DATA_BLOCK "PanelTorreCav"   // DB21
{ S7_Optimized_Access := 'FALSE' }
VERSION : 0.1
   VAR
      InhMV030 : Bool;   // Inhibición MV030
      InhMV031 : Bool;   // Inhibición MV031
      InhMP014 : Bool;   // Inhibición MP014
      InhMP015 : Bool;   // Inhibición MP015
      Flanco1MV030 : Bool;   // Flanco 1 MV030
      Flanco1MV031 : Bool;   // Flanco 1 MV031
      Flanco1MP014 : Bool;   // Flanco 1 MP014
      Flanco1MP015 : Bool;   // Flanco 1 MP015
      Flanco2MV030 : Bool;   // Flanco 2 MV030
      Flanco2MV031 : Bool;   // Flanco 2 MV031
      Flanco2MP014 : Bool;   // Flanco 2 MP014
      Flanco2MP015 : Bool;   // Flanco 2 MP015
      Flanco3MV030 : Bool;   // Flanco 3 MV030
      Flanco3MV031 : Bool;   // Flanco 3 MV031
      Flanco3MP014 : Bool;   // Flanco 3 MP014
      Flanco3MP015 : Bool;   // Flanco 3 MP015
      HabPanelMV030 : Bool;   // Habilitación desde Panel MV030
      HabPanelMV031 : Bool;   // Habilitación desde Panel MV031
      HabPanelMP014 : Bool;   // Habilitación desde Panel MP014
      HabPanelMP015 : Bool;   // Habilitación desde Panel MP015
      DeshabPanelMV030 : Bool;   // Deshabilitación desde Panel MV030
      DeshabPanelMV031 : Bool;   // Deshabilitación desde Panel MV031
      DeshabPanelMP014 : Bool;   // Deshabilitación desde Panel MP014
      DeshabPanelMP015 : Bool;   // Deshabilitación desde Panel MP015
      MarchaPanelMV030 : Bool;   // Marcha desde Panel MV030
      MarchaPanelMV031 : Bool;   // Marcha desde Panel MV031
      MarchaPanelMP014 : Bool;   // Marcha desde Panel MP014
      MarchaPanelMP015 : Bool;   // Marcha desde Panel MP015
      ParadaPanelMV030 : Bool;   // Parada desde Panel MV030
      ParadaPanelMV031 : Bool;   // Parada desde Panel MV031
      ParadaPanelMP014 : Bool;   // Parada desde Panel MP014
      ParadaPanelMP015 : Bool;   // Parada desde Panel MP015
      HabMV030 : Bool;   // Habilitado MV030
      HabMV031 : Bool;   // Habilitado MV031
      HabMP014 : Bool;   // Habilitado MP014
      HabMP015 : Bool;   // Habilitado MP015
      DeshabMV030 : Bool;   // Deshabilitado MV030
      DeshabMV031 : Bool;   // Deshabilitado MV031
      DeshabMP014 : Bool;   // Deshabilitado MP014
      DeshabMP015 : Bool;   // Deshabilitado MP015
      MarchaMV030 : Bool;   // Marchando MV030
      MarchaMV031 : Bool;   // Marchando MV031
      MarchaMP014 : Bool;   // Marchando MP014
      MarchaMP015 : Bool;   // Marchando MP015
      ParadaMV030 : Bool;   // Parando MV030
      ParadaMV031 : Bool;   // Parando MV031
      ParadaMP014 : Bool;   // Parando MP014
      ParadaMP015 : Bool;   // Parando MP015
      MantMV030 : Bool;   // Mantenimiento MV030
      MantMV031 : Bool;   // Mantenimiento MV031
      MantMP014 : Bool;   // Mantenimiento MP014
      MantMP015 : Bool;   // Mantenimiento MP015
      AutoV030 : Bool;   // Ventilador Controlado por temperatura V030
      AutoV031 : Bool;   // Ventilador Controlado por temperatura V031
      SPonV030 : Int;   // Setpoint arranque para V001
      SPonV031 : Int;   // Setpoint arranque para V002
      SPoffV030 : Int;   // Setpoint parada para V001
      SPoffV031 : Int;   // Setpoint parada para V002
      Temperatura : Int;   // Temperatura agua de torres
      ArranqueAutoV030 : Bool;   // Arranque Automático de ventilador 1
      ArranqueAutoV031 : Bool;   // Arranque Automático de ventilador 2
      Reserva_13 : Bool;
      Reserva_14 : Bool;
      Reserva_15 : Bool;
      Reserva_16 : Bool;
      Reserva_17 : Bool;
      Reserva_18 : Bool;
      Reserva_19 : Bool;
      Reserva_110 : Bool;
      Reserva_111 : Bool;
      Reserva_112 : Bool;
      Reserva_113 : Bool;
      Reserva_114 : Bool;
      Reserva_115 : Bool;
      Reserva_116 : Bool;
      Reserva_117 : Bool;
      Reserva_118 : Bool;
      Reserva_119 : Bool;
      Reserva_120 : Bool;
      Reserva_121 : Bool;
      Reserva_122 : Bool;
      Reserva_123 : Bool;
      Reserva_124 : Bool;
      Reserva_125 : Bool;
      Reserva_126 : Bool;
      Reserva_127 : Bool;
      Reserva_128 : Bool;
      Reserva_129 : Bool;
      Reserva_130 : Bool;
      Reserva_131 : Bool;
      Reserva_132 : Bool;
      Reserva_133 : Bool;
      Reserva_134 : Bool;
      Reserva_135 : Bool;
      Reserva_136 : Bool;
      Reserva_137 : Bool;
      Reserva_138 : Bool;
      Reserva_139 : Bool;
      Reserva_140 : Bool;
      Reserva_141 : Bool;
      Reserva_142 : Bool;
      Reserva_143 : Bool;
   END_VAR
BEGIN
END_DATA_BLOCK

DATA_BLOCK "TAguaCAV"   // DB51
{ S7_Optimized_Access := 'FALSE' }
AUTHOR : AEB
VERSION : 0.1
   VAR
      PrAlta : Real := 3.585069e+1;   // Presión Aire de Alta
      TmpCav : Real := 2.061632e+1;   // Temp Torre Cavaleto
      PrAlta2 : Real := 3.541667e+1;   // Presión Aire de Alta_Redundante
      PrBaja : Real := 6.140046e+0;   // Presión Aire de Baja
      STAT4 : Real;
      STAT5 : Real;
      STAT6 : Real;
      STAT7 : Real;
      STAT8 : Real;
      STAT9 : Real;
      STAT10 : Real := 1.446759e-3;
      STAT11 : Real;
      STAT12 : Real;
      STAT13 : Real;
      STAT14 : Real;
      STAT15 : Real;
      STAT16 : Real;
      STAT17 : Real;
      STAT18 : Real;
      STAT19 : Real;
      STAT20 : Real;
      STAT21 : Real;
      STAT22 : Real;
      STAT23 : Real;
      STAT24 : Real;
      STAT25 : Real;
      STAT26 : Real;
      STAT27 : Real;
      STAT28 : Real;
      STAT29 : Real;
      STAT30 : Real;
      STAT31 : Real;
      STAT32 : Real;
      STAT33 : Real;
      STAT34 : Real;
      STAT35 : Real;
      STAT36 : Real;
      STAT37 : Real;
      STAT38 : Real;
      STAT39 : Real;
      STAT40 : Real;
      STAT41 : Real;
      STAT42 : Real;
      STAT43 : Real;
      STAT44 : Real;
      STAT45 : Real;
      STAT46 : Real;
      STAT47 : Real;
      STAT48 : Real;
      STAT49 : Real;
      STAT50 : Real;
      STAT51 : Real;
      STAT52 : Real;
      STAT53 : Real;
      STAT54 : Real;
      STAT55 : Real;
      STAT56 : Real;
      STAT57 : Real;
      STAT58 : Real;
      STAT59 : Real;
      STAT60 : Real;
      STAT61 : Real;
      STAT62 : Real;
      STAT63 : Real;
      STAT64 : Real;
      STAT65 : Real;
   END_VAR
BEGIN
END_DATA_BLOCK

// folder: Torres de Agua/Torres Chillers

DATA_BLOCK "CFG-TorresCH"   // DB92
{ S7_Optimized_Access := 'FALSE' }
VERSION : 0.1
   VAR
      AutoV001 : Bool;   // Ventilador Controlado por temperatura V001
      AutoV002 : Bool;   // Ventilador Controlado por temperatura V002
      AutoV003 : Bool;   // Ventilador Controlado por temperatura V003
      SPonV001 : Int;   // Setpoint arranque para V001
      SPonV002 : Int;   // Setpoint arranque para V002
      SPonV003 : Int;   // Setpoint arranque para V003
      SPoffV001 : Int;   // Setpoint parada para V001
      SPoffV002 : Int;   // Setpoint parada para V002
      SPoffV003 : Int;   // Setpoint parada para V003
      Temperatura : Int;   // Temperatura agua de torres
      ArranqueAutoV001 : Bool;   // Arranque Automático de ventilador 1
      ArranqueAutoV002 : Bool;   // Arranque Automático de ventilador 2
      ArranqueAutoV003 : Bool;   // Arranque Automático de ventilador 3
   END_VAR
BEGIN
END_DATA_BLOCK

// folder: (top level)

FUNCTION "Arranques General" : Void   // FC4, LAD
{ S7_Optimized_Access := 'FALSE' }
VERSION : 0.1
   VAR_TEMP
      TEMP0 : Bool;
      TEMP1 : Bool;
      TEMP2 : Bool;
      TEMP3 : Bool;
      TEMP4 : Bool;
   END_VAR
   VAR_TEMP   // added for the SCL form of the ladder/FBD networks
      _w1 : Bool;
      _w2 : Bool;
      _s5time1 : S5Time;
   END_VAR
BEGIN

REGION Network 1: Motor MT007 - Bomba Soplado L1 / Bloque motor MT007 - Bomba Soplado L1
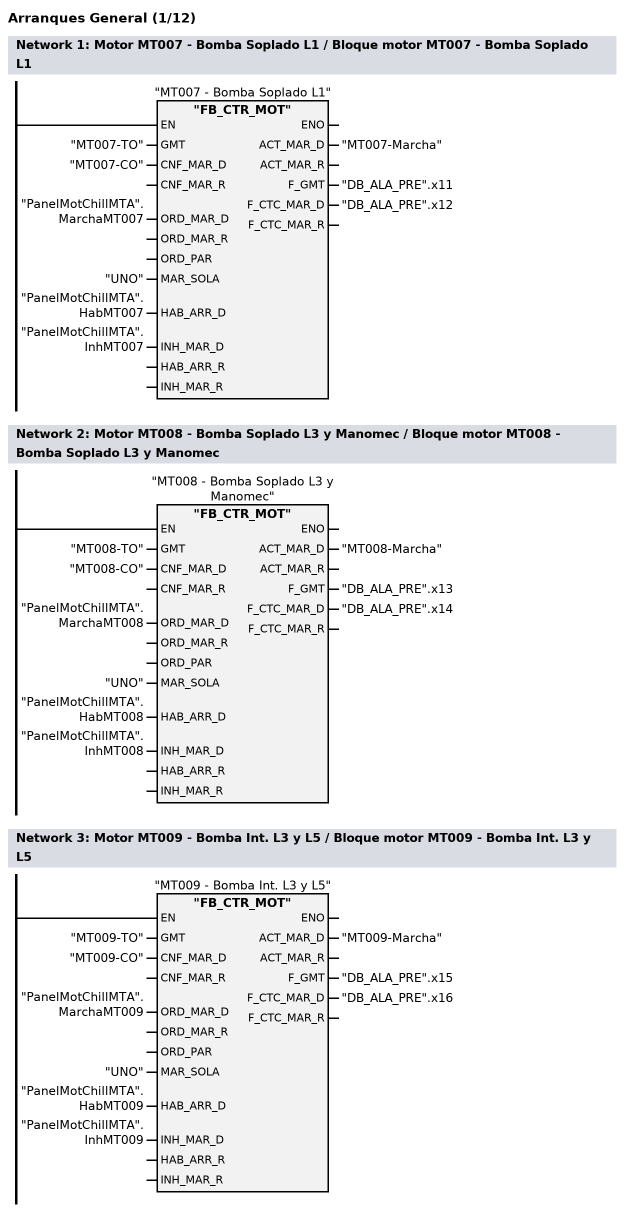
   RUNG wire#powerrail
      "MT007 - Bomba Soplado L1"(GMT := "MT007-TO", CNF_MAR_D := "MT007-CO", CNF_MAR_R :=, ORD_MAR_D := "PanelMotChillMTA".MarchaMT007, ORD_MAR_R :=, ORD_PAR :=, MAR_SOLA := "UNO", HAB_ARR_D := "PanelMotChillMTA".HabMT007, INH_MAR_D := "PanelMotChillMTA".InhMT007, HAB_ARR_R :=, INH_MAR_R :=, ACT_MAR_D => "MT007-Marcha", ACT_MAR_R =>, F_GMT => "DB_ALA_PRE".x11, F_CTC_MAR_D => "DB_ALA_PRE".x12, F_CTC_MAR_R =>)
   END_RUNG
   // the same network as SCL:
   "MT007 - Bomba Soplado L1"(GMT := "MT007-TO",   // "FB_CTR_MOT"
                           CNF_MAR_D := "MT007-CO",
                           ORD_MAR_D := "PanelMotChillMTA".MarchaMT007,
                           MAR_SOLA := "UNO",
                           HAB_ARR_D := "PanelMotChillMTA".HabMT007,
                           INH_MAR_D := "PanelMotChillMTA".InhMT007,
                           ACT_MAR_D => "MT007-Marcha",
                           F_GMT => "DB_ALA_PRE".x11,
                           F_CTC_MAR_D => "DB_ALA_PRE".x12);
END_REGION

REGION Network 2: Motor MT008 - Bomba Soplado L3 y Manomec / Bloque motor MT008 - Bomba Soplado L3 y Manomec
   RUNG wire#powerrail
      "MT008 - Bomba Soplado L3 y Manomec"(GMT := "MT008-TO", CNF_MAR_D := "MT008-CO", CNF_MAR_R :=, ORD_MAR_D := "PanelMotChillMTA".MarchaMT008, ORD_MAR_R :=, ORD_PAR :=, MAR_SOLA := "UNO", HAB_ARR_D := "PanelMotChillMTA".HabMT008, INH_MAR_D := "PanelMotChillMTA".InhMT008, HAB_ARR_R :=, INH_MAR_R :=, ACT_MAR_D => "MT008-Marcha", ACT_MAR_R =>, F_GMT => "DB_ALA_PRE".x13, F_CTC_MAR_D => "DB_ALA_PRE".x14, F_CTC_MAR_R =>)
   END_RUNG
   // the same network as SCL:
   "MT008 - Bomba Soplado L3 y Manomec"(GMT := "MT008-TO",   // "FB_CTR_MOT"
                           CNF_MAR_D := "MT008-CO",
                           ORD_MAR_D := "PanelMotChillMTA".MarchaMT008,
                           MAR_SOLA := "UNO",
                           HAB_ARR_D := "PanelMotChillMTA".HabMT008,
                           INH_MAR_D := "PanelMotChillMTA".InhMT008,
                           ACT_MAR_D => "MT008-Marcha",
                           F_GMT => "DB_ALA_PRE".x13,
                           F_CTC_MAR_D => "DB_ALA_PRE".x14);
END_REGION

REGION Network 3: Motor MT009 - Bomba Int. L3 y L5 / Bloque motor MT009 - Bomba Int. L3 y L5
   RUNG wire#powerrail
      "MT009 - Bomba Int. L3 y L5"(GMT := "MT009-TO", CNF_MAR_D := "MT009-CO", CNF_MAR_R :=, ORD_MAR_D := "PanelMotChillMTA".MarchaMT009, ORD_MAR_R :=, ORD_PAR :=, MAR_SOLA := "UNO", HAB_ARR_D := "PanelMotChillMTA".HabMT009, INH_MAR_D := "PanelMotChillMTA".InhMT009, HAB_ARR_R :=, INH_MAR_R :=, ACT_MAR_D => "MT009-Marcha", ACT_MAR_R =>, F_GMT => "DB_ALA_PRE".x15, F_CTC_MAR_D => "DB_ALA_PRE".x16, F_CTC_MAR_R =>)
   END_RUNG
   // the same network as SCL:
   "MT009 - Bomba Int. L3 y L5"(GMT := "MT009-TO",   // "FB_CTR_MOT"
                           CNF_MAR_D := "MT009-CO",
                           ORD_MAR_D := "PanelMotChillMTA".MarchaMT009,
                           MAR_SOLA := "UNO",
                           HAB_ARR_D := "PanelMotChillMTA".HabMT009,
                           INH_MAR_D := "PanelMotChillMTA".InhMT009,
                           ACT_MAR_D => "MT009-Marcha",
                           F_GMT => "DB_ALA_PRE".x15,
                           F_CTC_MAR_D => "DB_ALA_PRE".x16);
END_REGION

REGION Network 4: Motor MT010 - Bomba Int L1 y Manomec / Bloque motor MT010 - Bomba Int L1 y Manomec
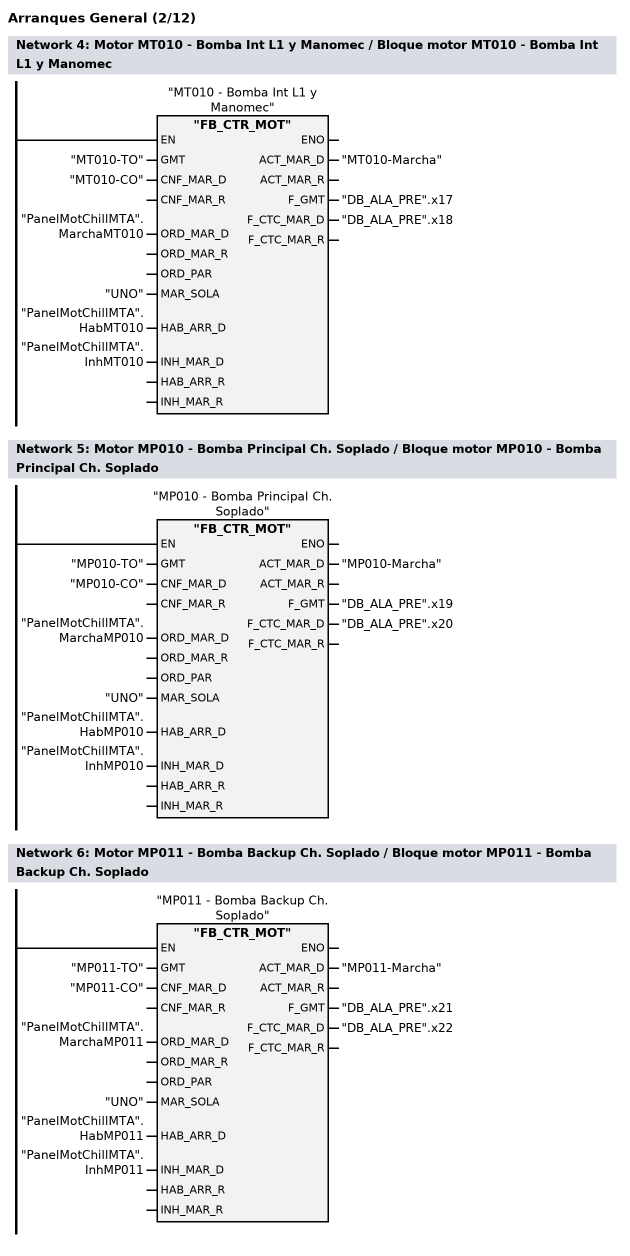
   RUNG wire#powerrail
      "MT010 - Bomba Int L1 y Manomec"(GMT := "MT010-TO", CNF_MAR_D := "MT010-CO", CNF_MAR_R :=, ORD_MAR_D := "PanelMotChillMTA".MarchaMT010, ORD_MAR_R :=, ORD_PAR :=, MAR_SOLA := "UNO", HAB_ARR_D := "PanelMotChillMTA".HabMT010, INH_MAR_D := "PanelMotChillMTA".InhMT010, HAB_ARR_R :=, INH_MAR_R :=, ACT_MAR_D => "MT010-Marcha", ACT_MAR_R =>, F_GMT => "DB_ALA_PRE".x17, F_CTC_MAR_D => "DB_ALA_PRE".x18, F_CTC_MAR_R =>)
   END_RUNG
   // the same network as SCL:
   "MT010 - Bomba Int L1 y Manomec"(GMT := "MT010-TO",   // "FB_CTR_MOT"
                           CNF_MAR_D := "MT010-CO",
                           ORD_MAR_D := "PanelMotChillMTA".MarchaMT010,
                           MAR_SOLA := "UNO",
                           HAB_ARR_D := "PanelMotChillMTA".HabMT010,
                           INH_MAR_D := "PanelMotChillMTA".InhMT010,
                           ACT_MAR_D => "MT010-Marcha",
                           F_GMT => "DB_ALA_PRE".x17,
                           F_CTC_MAR_D => "DB_ALA_PRE".x18);
END_REGION

REGION Network 5: Motor MP010 - Bomba Principal Ch. Soplado / Bloque motor MP010 - Bomba Principal Ch. Soplado
   RUNG wire#powerrail
      "MP010 - Bomba Principal Ch. Soplado"(GMT := "MP010-TO", CNF_MAR_D := "MP010-CO", CNF_MAR_R :=, ORD_MAR_D := "PanelMotChillMTA".MarchaMP010, ORD_MAR_R :=, ORD_PAR :=, MAR_SOLA := "UNO", HAB_ARR_D := "PanelMotChillMTA".HabMP010, INH_MAR_D := "PanelMotChillMTA".InhMP010, HAB_ARR_R :=, INH_MAR_R :=, ACT_MAR_D => "MP010-Marcha", ACT_MAR_R =>, F_GMT => "DB_ALA_PRE".x19, F_CTC_MAR_D => "DB_ALA_PRE".x20, F_CTC_MAR_R =>)
   END_RUNG
   // the same network as SCL:
   "MP010 - Bomba Principal Ch. Soplado"(GMT := "MP010-TO",   // "FB_CTR_MOT"
                           CNF_MAR_D := "MP010-CO",
                           ORD_MAR_D := "PanelMotChillMTA".MarchaMP010,
                           MAR_SOLA := "UNO",
                           HAB_ARR_D := "PanelMotChillMTA".HabMP010,
                           INH_MAR_D := "PanelMotChillMTA".InhMP010,
                           ACT_MAR_D => "MP010-Marcha",
                           F_GMT => "DB_ALA_PRE".x19,
                           F_CTC_MAR_D => "DB_ALA_PRE".x20);
END_REGION

REGION Network 6: Motor MP011 - Bomba Backup Ch. Soplado / Bloque motor MP011 - Bomba Backup Ch. Soplado
   RUNG wire#powerrail
      "MP011 - Bomba Backup Ch. Soplado"(GMT := "MP011-TO", CNF_MAR_D := "MP011-CO", CNF_MAR_R :=, ORD_MAR_D := "PanelMotChillMTA".MarchaMP011, ORD_MAR_R :=, ORD_PAR :=, MAR_SOLA := "UNO", HAB_ARR_D := "PanelMotChillMTA".HabMP011, INH_MAR_D := "PanelMotChillMTA".InhMP011, HAB_ARR_R :=, INH_MAR_R :=, ACT_MAR_D => "MP011-Marcha", ACT_MAR_R =>, F_GMT => "DB_ALA_PRE".x21, F_CTC_MAR_D => "DB_ALA_PRE".x22, F_CTC_MAR_R =>)
   END_RUNG
   // the same network as SCL:
   "MP011 - Bomba Backup Ch. Soplado"(GMT := "MP011-TO",   // "FB_CTR_MOT"
                           CNF_MAR_D := "MP011-CO",
                           ORD_MAR_D := "PanelMotChillMTA".MarchaMP011,
                           MAR_SOLA := "UNO",
                           HAB_ARR_D := "PanelMotChillMTA".HabMP011,
                           INH_MAR_D := "PanelMotChillMTA".InhMP011,
                           ACT_MAR_D => "MP011-Marcha",
                           F_GMT => "DB_ALA_PRE".x21,
                           F_CTC_MAR_D => "DB_ALA_PRE".x22);
END_REGION

REGION Network 7: Motor MP012 - Bomba Principal Ch. Envasado / Bloque motor MP012 - Bomba Principal Ch. Envasado
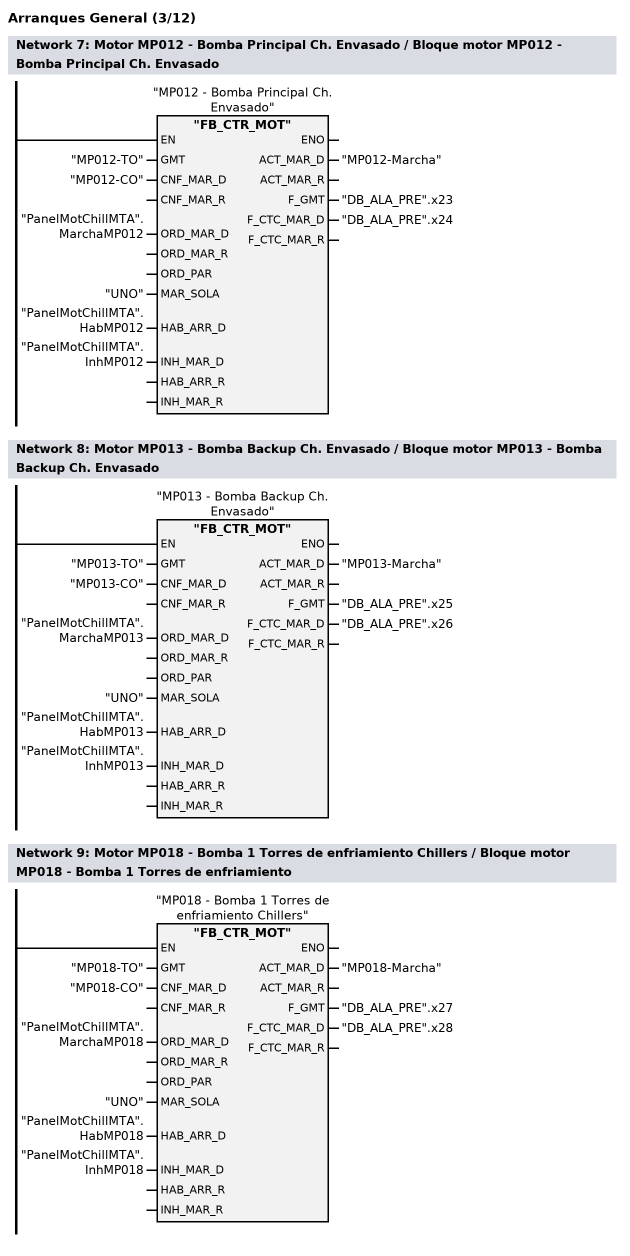
   RUNG wire#powerrail
      "MP012 - Bomba Principal Ch. Envasado"(GMT := "MP012-TO", CNF_MAR_D := "MP012-CO", CNF_MAR_R :=, ORD_MAR_D := "PanelMotChillMTA".MarchaMP012, ORD_MAR_R :=, ORD_PAR :=, MAR_SOLA := "UNO", HAB_ARR_D := "PanelMotChillMTA".HabMP012, INH_MAR_D := "PanelMotChillMTA".InhMP012, HAB_ARR_R :=, INH_MAR_R :=, ACT_MAR_D => "MP012-Marcha", ACT_MAR_R =>, F_GMT => "DB_ALA_PRE".x23, F_CTC_MAR_D => "DB_ALA_PRE".x24, F_CTC_MAR_R =>)
   END_RUNG
   // the same network as SCL:
   "MP012 - Bomba Principal Ch. Envasado"(GMT := "MP012-TO",   // "FB_CTR_MOT"
                           CNF_MAR_D := "MP012-CO",
                           ORD_MAR_D := "PanelMotChillMTA".MarchaMP012,
                           MAR_SOLA := "UNO",
                           HAB_ARR_D := "PanelMotChillMTA".HabMP012,
                           INH_MAR_D := "PanelMotChillMTA".InhMP012,
                           ACT_MAR_D => "MP012-Marcha",
                           F_GMT => "DB_ALA_PRE".x23,
                           F_CTC_MAR_D => "DB_ALA_PRE".x24);
END_REGION

REGION Network 8: Motor MP013 - Bomba Backup Ch. Envasado / Bloque motor MP013 - Bomba Backup Ch. Envasado
   RUNG wire#powerrail
      "MP013 - Bomba Backup Ch. Envasado"(GMT := "MP013-TO", CNF_MAR_D := "MP013-CO", CNF_MAR_R :=, ORD_MAR_D := "PanelMotChillMTA".MarchaMP013, ORD_MAR_R :=, ORD_PAR :=, MAR_SOLA := "UNO", HAB_ARR_D := "PanelMotChillMTA".HabMP013, INH_MAR_D := "PanelMotChillMTA".InhMP013, HAB_ARR_R :=, INH_MAR_R :=, ACT_MAR_D => "MP013-Marcha", ACT_MAR_R =>, F_GMT => "DB_ALA_PRE".x25, F_CTC_MAR_D => "DB_ALA_PRE".x26, F_CTC_MAR_R =>)
   END_RUNG
   // the same network as SCL:
   "MP013 - Bomba Backup Ch. Envasado"(GMT := "MP013-TO",   // "FB_CTR_MOT"
                           CNF_MAR_D := "MP013-CO",
                           ORD_MAR_D := "PanelMotChillMTA".MarchaMP013,
                           MAR_SOLA := "UNO",
                           HAB_ARR_D := "PanelMotChillMTA".HabMP013,
                           INH_MAR_D := "PanelMotChillMTA".InhMP013,
                           ACT_MAR_D => "MP013-Marcha",
                           F_GMT => "DB_ALA_PRE".x25,
                           F_CTC_MAR_D => "DB_ALA_PRE".x26);
END_REGION

REGION Network 9: Motor MP018 - Bomba 1 Torres de enfriamiento Chillers / Bloque motor MP018 - Bomba 1 Torres de enfriamiento
   RUNG wire#powerrail
      "MP018 - Bomba 1 Torres de enfriamiento Chillers"(GMT := "MP018-TO", CNF_MAR_D := "MP018-CO", CNF_MAR_R :=, ORD_MAR_D := "PanelMotChillMTA".MarchaMP018, ORD_MAR_R :=, ORD_PAR :=, MAR_SOLA := "UNO", HAB_ARR_D := "PanelMotChillMTA".HabMP018, INH_MAR_D := "PanelMotChillMTA".InhMP018, HAB_ARR_R :=, INH_MAR_R :=, ACT_MAR_D => "MP018-Marcha", ACT_MAR_R =>, F_GMT => "DB_ALA_PRE".x27, F_CTC_MAR_D => "DB_ALA_PRE".x28, F_CTC_MAR_R =>)
   END_RUNG
   // the same network as SCL:
   "MP018 - Bomba 1 Torres de enfriamiento Chillers"(GMT := "MP018-TO",   // "FB_CTR_MOT"
                           CNF_MAR_D := "MP018-CO",
                           ORD_MAR_D := "PanelMotChillMTA".MarchaMP018,
                           MAR_SOLA := "UNO",
                           HAB_ARR_D := "PanelMotChillMTA".HabMP018,
                           INH_MAR_D := "PanelMotChillMTA".InhMP018,
                           ACT_MAR_D => "MP018-Marcha",
                           F_GMT => "DB_ALA_PRE".x27,
                           F_CTC_MAR_D => "DB_ALA_PRE".x28);
END_REGION

REGION Network 10: Motor MP019 - Bomba 2 Torres de enfriamiento Chillers / Bloque motor MP019 - Bomba 2 Torres de enfriamiento
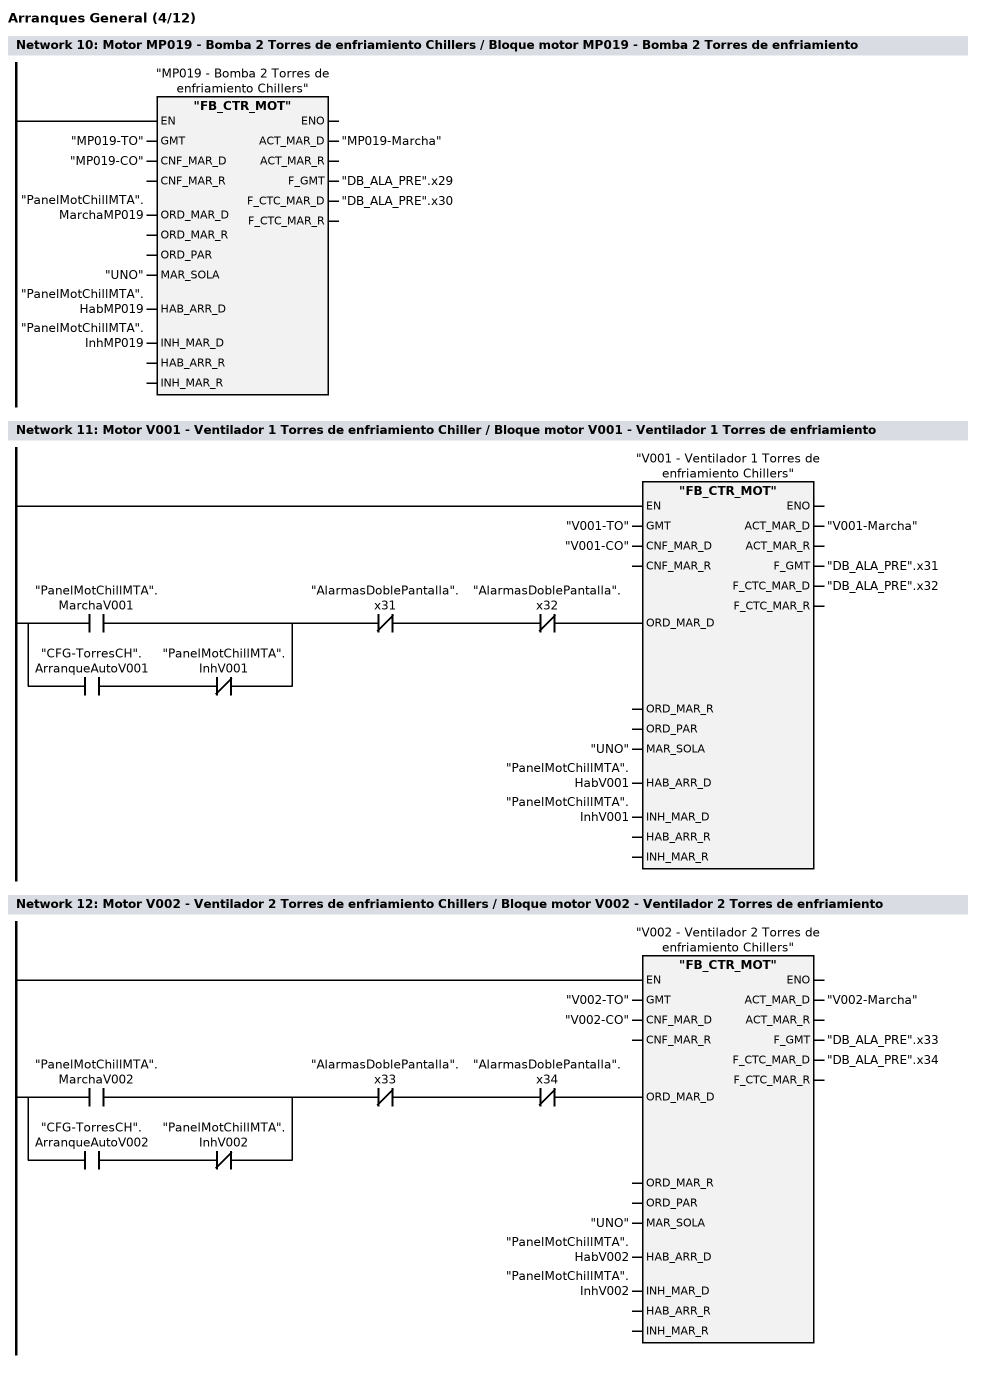
   RUNG wire#powerrail
      "MP019 - Bomba 2 Torres de enfriamiento Chillers"(GMT := "MP019-TO", CNF_MAR_D := "MP019-CO", CNF_MAR_R :=, ORD_MAR_D := "PanelMotChillMTA".MarchaMP019, ORD_MAR_R :=, ORD_PAR :=, MAR_SOLA := "UNO", HAB_ARR_D := "PanelMotChillMTA".HabMP019, INH_MAR_D := "PanelMotChillMTA".InhMP019, HAB_ARR_R :=, INH_MAR_R :=, ACT_MAR_D => "MP019-Marcha", ACT_MAR_R =>, F_GMT => "DB_ALA_PRE".x29, F_CTC_MAR_D => "DB_ALA_PRE".x30, F_CTC_MAR_R =>)
   END_RUNG
   // the same network as SCL:
   "MP019 - Bomba 2 Torres de enfriamiento Chillers"(GMT := "MP019-TO",   // "FB_CTR_MOT"
                           CNF_MAR_D := "MP019-CO",
                           ORD_MAR_D := "PanelMotChillMTA".MarchaMP019,
                           MAR_SOLA := "UNO",
                           HAB_ARR_D := "PanelMotChillMTA".HabMP019,
                           INH_MAR_D := "PanelMotChillMTA".InhMP019,
                           ACT_MAR_D => "MP019-Marcha",
                           F_GMT => "DB_ALA_PRE".x29,
                           F_CTC_MAR_D => "DB_ALA_PRE".x30);
END_REGION

REGION Network 11: Motor V001 - Ventilador 1 Torres de enfriamiento Chiller / Bloque motor V001 - Ventilador 1 Torres de enfriamiento
   RUNG wire#powerrail
      "V001 - Ventilador 1 Torres de enfriamiento Chillers"(ORD_MAR_D := wire#w2, GMT := "V001-TO", CNF_MAR_D := "V001-CO", CNF_MAR_R :=, ORD_MAR_R :=, ORD_PAR :=, MAR_SOLA := "UNO", HAB_ARR_D := "PanelMotChillMTA".HabV001, INH_MAR_D := "PanelMotChillMTA".InhV001, HAB_ARR_R :=, INH_MAR_R :=, ACT_MAR_D => "V001-Marcha", ACT_MAR_R =>, F_GMT => "DB_ALA_PRE".x31, F_CTC_MAR_D => "DB_ALA_PRE".x32, F_CTC_MAR_R =>)
   END_RUNG
   RUNG wire#powerrail
      Contact( "PanelMotChillMTA".MarchaV001 )
      wire#w1
      I_Contact( "AlarmasDoblePantalla".x31 )
      I_Contact( "AlarmasDoblePantalla".x32 )
   END_RUNG wire#w2
   RUNG wire#powerrail
      Contact( "CFG-TorresCH".ArranqueAutoV001 )
      I_Contact( "PanelMotChillMTA".InhV001 )
   END_RUNG wire#w1
   // the same network as SCL:
   "V001 - Ventilador 1 Torres de enfriamiento Chillers"(GMT := "V001-TO",   // "FB_CTR_MOT"
                           CNF_MAR_D := "V001-CO",
                           ORD_MAR_D := ("PanelMotChillMTA".MarchaV001 OR ("CFG-TorresCH".ArranqueAutoV001 AND NOT "PanelMotChillMTA".InhV001)) AND NOT "AlarmasDoblePantalla".x31 AND NOT "AlarmasDoblePantalla".x32,
                           MAR_SOLA := "UNO",
                           HAB_ARR_D := "PanelMotChillMTA".HabV001,
                           INH_MAR_D := "PanelMotChillMTA".InhV001,
                           ACT_MAR_D => "V001-Marcha",
                           F_GMT => "DB_ALA_PRE".x31,
                           F_CTC_MAR_D => "DB_ALA_PRE".x32);
END_REGION

REGION Network 12: Motor V002 - Ventilador 2 Torres de enfriamiento Chillers / Bloque motor V002 - Ventilador 2 Torres de enfriamiento
   RUNG wire#powerrail
      "V002 - Ventilador 2 Torres de enfriamiento Chillers"(ORD_MAR_D := wire#w2, GMT := "V002-TO", CNF_MAR_D := "V002-CO", CNF_MAR_R :=, ORD_MAR_R :=, ORD_PAR :=, MAR_SOLA := "UNO", HAB_ARR_D := "PanelMotChillMTA".HabV002, INH_MAR_D := "PanelMotChillMTA".InhV002, HAB_ARR_R :=, INH_MAR_R :=, ACT_MAR_D => "V002-Marcha", ACT_MAR_R =>, F_GMT => "DB_ALA_PRE".x33, F_CTC_MAR_D => "DB_ALA_PRE".x34, F_CTC_MAR_R =>)
   END_RUNG
   RUNG wire#powerrail
      Contact( "PanelMotChillMTA".MarchaV002 )
      wire#w1
      I_Contact( "AlarmasDoblePantalla".x33 )
      I_Contact( "AlarmasDoblePantalla".x34 )
   END_RUNG wire#w2
   RUNG wire#powerrail
      Contact( "CFG-TorresCH".ArranqueAutoV002 )
      I_Contact( "PanelMotChillMTA".InhV002 )
   END_RUNG wire#w1
   // the same network as SCL:
   "V002 - Ventilador 2 Torres de enfriamiento Chillers"(GMT := "V002-TO",   // "FB_CTR_MOT"
                           CNF_MAR_D := "V002-CO",
                           ORD_MAR_D := ("PanelMotChillMTA".MarchaV002 OR ("CFG-TorresCH".ArranqueAutoV002 AND NOT "PanelMotChillMTA".InhV002)) AND NOT "AlarmasDoblePantalla".x33 AND NOT "AlarmasDoblePantalla".x34,
                           MAR_SOLA := "UNO",
                           HAB_ARR_D := "PanelMotChillMTA".HabV002,
                           INH_MAR_D := "PanelMotChillMTA".InhV002,
                           ACT_MAR_D => "V002-Marcha",
                           F_GMT => "DB_ALA_PRE".x33,
                           F_CTC_MAR_D => "DB_ALA_PRE".x34);
END_REGION

REGION Network 13: Motor V003 - Ventilador 3 Torres de enfriamiento Chillers / Bloque motor V003 - Ventilador 3 Torres de enfriamiento
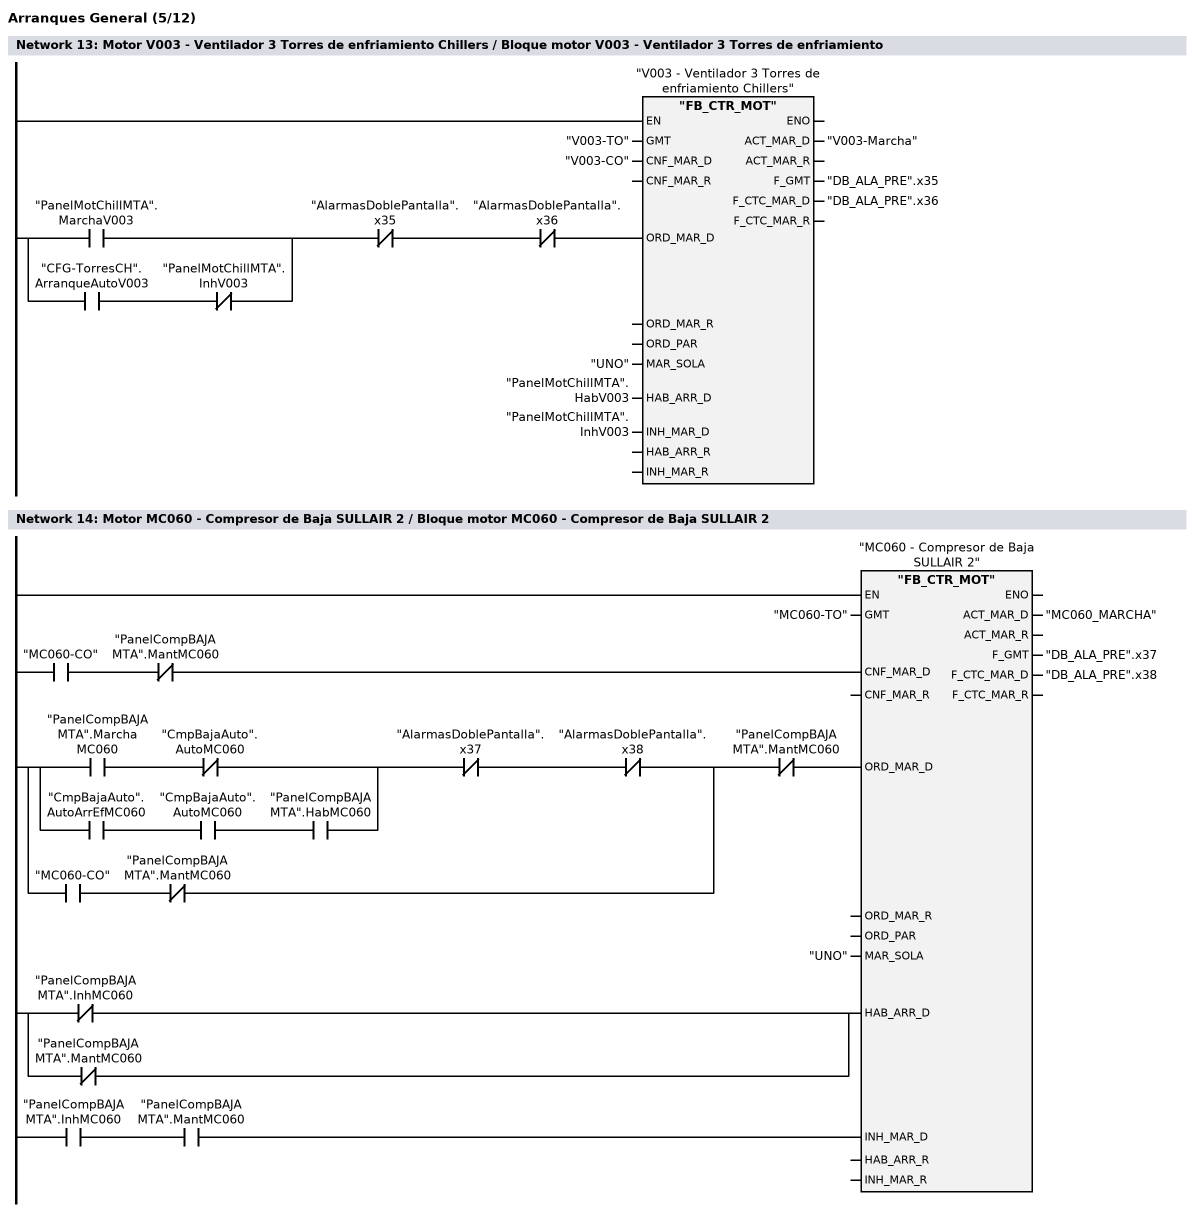
   RUNG wire#powerrail
      "V003 - Ventilador 3 Torres de enfriamiento Chillers"(ORD_MAR_D := wire#w2, GMT := "V003-TO", CNF_MAR_D := "V003-CO", CNF_MAR_R :=, ORD_MAR_R :=, ORD_PAR :=, MAR_SOLA := "UNO", HAB_ARR_D := "PanelMotChillMTA".HabV003, INH_MAR_D := "PanelMotChillMTA".InhV003, HAB_ARR_R :=, INH_MAR_R :=, ACT_MAR_D => "V003-Marcha", ACT_MAR_R =>, F_GMT => "DB_ALA_PRE".x35, F_CTC_MAR_D => "DB_ALA_PRE".x36, F_CTC_MAR_R =>)
   END_RUNG
   RUNG wire#powerrail
      Contact( "PanelMotChillMTA".MarchaV003 )
      wire#w1
      I_Contact( "AlarmasDoblePantalla".x35 )
      I_Contact( "AlarmasDoblePantalla".x36 )
   END_RUNG wire#w2
   RUNG wire#powerrail
      Contact( "CFG-TorresCH".ArranqueAutoV003 )
      I_Contact( "PanelMotChillMTA".InhV003 )
   END_RUNG wire#w1
   // the same network as SCL:
   "V003 - Ventilador 3 Torres de enfriamiento Chillers"(GMT := "V003-TO",   // "FB_CTR_MOT"
                           CNF_MAR_D := "V003-CO",
                           ORD_MAR_D := ("PanelMotChillMTA".MarchaV003 OR ("CFG-TorresCH".ArranqueAutoV003 AND NOT "PanelMotChillMTA".InhV003)) AND NOT "AlarmasDoblePantalla".x35 AND NOT "AlarmasDoblePantalla".x36,
                           MAR_SOLA := "UNO",
                           HAB_ARR_D := "PanelMotChillMTA".HabV003,
                           INH_MAR_D := "PanelMotChillMTA".InhV003,
                           ACT_MAR_D => "V003-Marcha",
                           F_GMT => "DB_ALA_PRE".x35,
                           F_CTC_MAR_D => "DB_ALA_PRE".x36);
END_REGION

REGION Network 14: Motor MC060 - Compresor de Baja SULLAIR 2 / Bloque motor MC060 - Compresor de Baja SULLAIR 2
   RUNG wire#powerrail
      "MC060 - Compresor de Baja SULLAIR 2"(CNF_MAR_D := wire#w1, ORD_MAR_D := wire#w4, HAB_ARR_D := wire#w5, INH_MAR_D := wire#w6, GMT := "MC060-TO", CNF_MAR_R :=, ORD_MAR_R :=, ORD_PAR :=, MAR_SOLA := "UNO", HAB_ARR_R :=, INH_MAR_R :=, ACT_MAR_D => "MC060_MARCHA", ACT_MAR_R =>, F_GMT => "DB_ALA_PRE".x37, F_CTC_MAR_D => "DB_ALA_PRE".x38, F_CTC_MAR_R =>)
   END_RUNG
   RUNG wire#powerrail
      Contact( "MC060-CO" )
      I_Contact( "PanelCompBAJA MTA".MantMC060 )
   END_RUNG wire#w1
   RUNG wire#powerrail
      Contact( "PanelCompBAJA MTA".MarchaMC060 )
      I_Contact( "CmpBajaAuto".AutoMC060 )
      wire#w2
      I_Contact( "AlarmasDoblePantalla".x37 )
      I_Contact( "AlarmasDoblePantalla".x38 )
      wire#w3
      I_Contact( "PanelCompBAJA MTA".MantMC060 )
   END_RUNG wire#w4
   RUNG wire#powerrail
      Contact( "CmpBajaAuto".AutoArrEfMC060 )
      Contact( "CmpBajaAuto".AutoMC060 )
      Contact( "PanelCompBAJA MTA".HabMC060 )
   END_RUNG wire#w2
   RUNG wire#powerrail
      Contact( "MC060-CO" )
      I_Contact( "PanelCompBAJA MTA".MantMC060 )
   END_RUNG wire#w3
   RUNG wire#powerrail
      I_Contact( "PanelCompBAJA MTA".InhMC060 )
   END_RUNG wire#w5
   RUNG wire#powerrail
      I_Contact( "PanelCompBAJA MTA".MantMC060 )
   END_RUNG wire#w5
   RUNG wire#powerrail
      Contact( "PanelCompBAJA MTA".InhMC060 )
      Contact( "PanelCompBAJA MTA".MantMC060 )
   END_RUNG wire#w6
   // the same network as SCL:
   "MC060 - Compresor de Baja SULLAIR 2"(GMT := "MC060-TO",   // "FB_CTR_MOT"
                           CNF_MAR_D := "MC060-CO" AND NOT "PanelCompBAJA MTA".MantMC060,
                           ORD_MAR_D := (((("PanelCompBAJA MTA".MarchaMC060 AND NOT "CmpBajaAuto".AutoMC060) OR ("CmpBajaAuto".AutoArrEfMC060 AND "CmpBajaAuto".AutoMC060 AND "PanelCompBAJA MTA".HabMC060)) AND NOT "AlarmasDoblePantalla".x37 AND NOT "AlarmasDoblePantalla".x38) OR ("MC060-CO" AND NOT "PanelCompBAJA MTA".MantMC060)) AND NOT "PanelCompBAJA MTA".MantMC060,
                           MAR_SOLA := "UNO",
                           HAB_ARR_D := NOT "PanelCompBAJA MTA".InhMC060 OR NOT "PanelCompBAJA MTA".MantMC060,
                           INH_MAR_D := "PanelCompBAJA MTA".InhMC060 AND "PanelCompBAJA MTA".MantMC060,
                           ACT_MAR_D => "MC060_MARCHA",
                           F_GMT => "DB_ALA_PRE".x37,
                           F_CTC_MAR_D => "DB_ALA_PRE".x38);
END_REGION

REGION Network 15
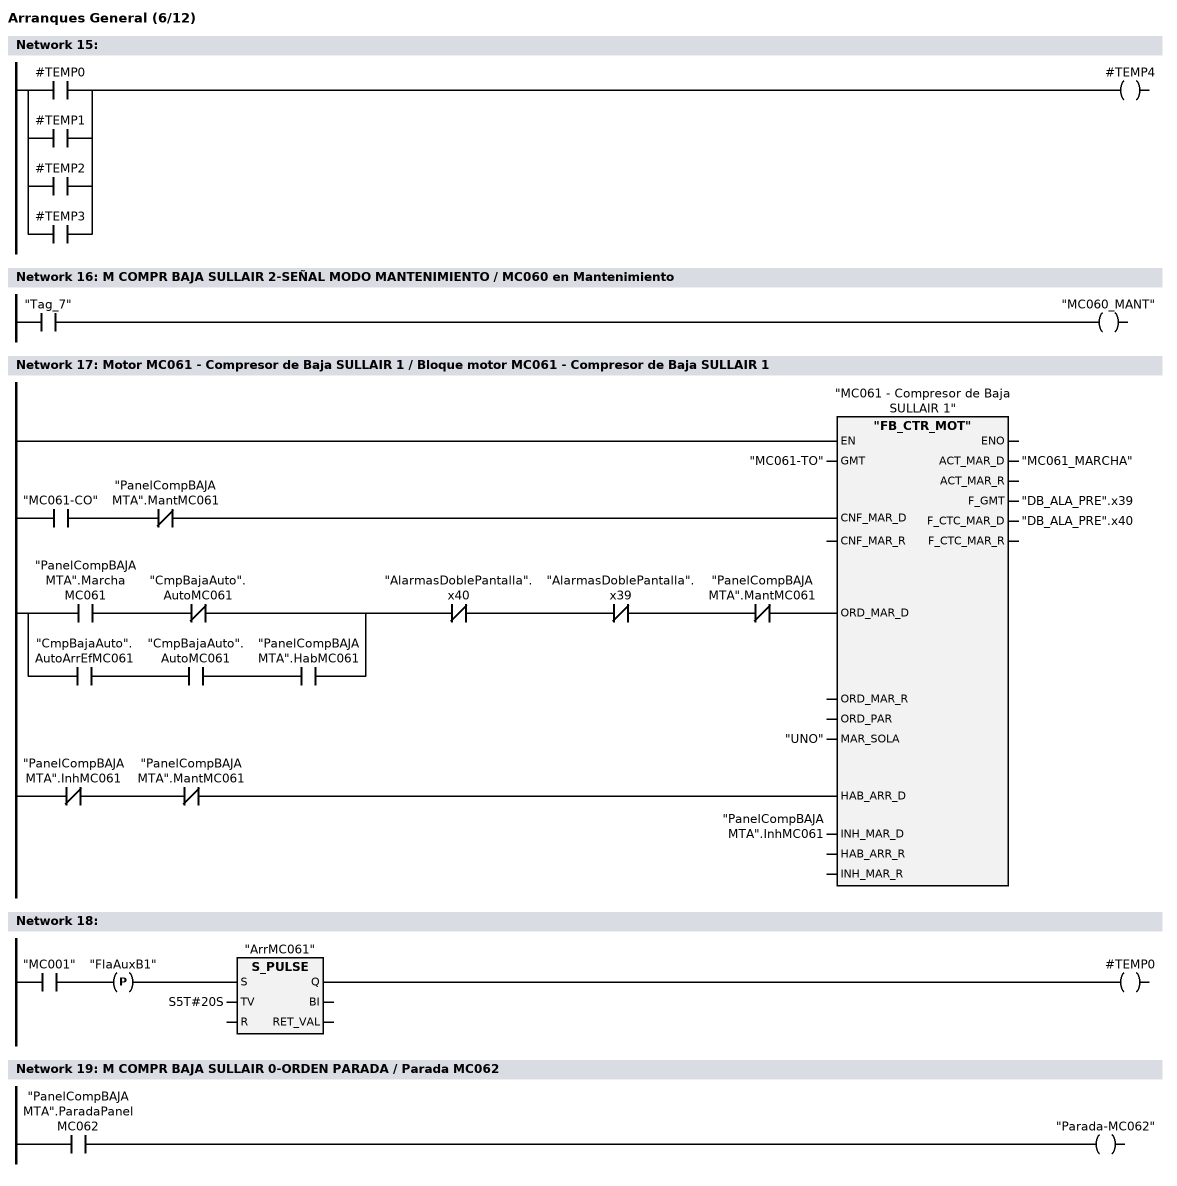
   RUNG wire#powerrail
      Contact( #TEMP0 )
      wire#w1
      Coil( #TEMP4 )
   END_RUNG
   RUNG wire#powerrail
      Contact( #TEMP1 )
   END_RUNG wire#w1
   RUNG wire#powerrail
      Contact( #TEMP2 )
   END_RUNG wire#w1
   RUNG wire#powerrail
      Contact( #TEMP3 )
   END_RUNG wire#w1
   // the same network as SCL:
   #TEMP4 := #TEMP0 OR #TEMP1 OR #TEMP2 OR #TEMP3;
END_REGION

REGION Network 16: M COMPR BAJA SULLAIR 2-SEÑAL MODO MANTENIMIENTO / MC060 en Mantenimiento
   RUNG wire#powerrail
      Contact( "Tag_7" )
      Coil( "MC060_MANT" )
   END_RUNG
   // the same network as SCL:
   "MC060_MANT" := "Tag_7";
END_REGION

REGION Network 17: Motor MC061 - Compresor de Baja SULLAIR 1 / Bloque motor MC061 - Compresor de Baja SULLAIR 1
   RUNG wire#powerrail
      "MC061 - Compresor de Baja SULLAIR 1"(CNF_MAR_D := wire#w1, ORD_MAR_D := wire#w3, HAB_ARR_D := wire#w4, GMT := "MC061-TO", CNF_MAR_R :=, ORD_MAR_R :=, ORD_PAR :=, MAR_SOLA := "UNO", INH_MAR_D := "PanelCompBAJA MTA".InhMC061, HAB_ARR_R :=, INH_MAR_R :=, ACT_MAR_D => "MC061_MARCHA", ACT_MAR_R =>, F_GMT => "DB_ALA_PRE".x39, F_CTC_MAR_D => "DB_ALA_PRE".x40, F_CTC_MAR_R =>)
   END_RUNG
   RUNG wire#powerrail
      Contact( "MC061-CO" )
      I_Contact( "PanelCompBAJA MTA".MantMC061 )
   END_RUNG wire#w1
   RUNG wire#powerrail
      Contact( "PanelCompBAJA MTA".MarchaMC061 )
      I_Contact( "CmpBajaAuto".AutoMC061 )
      wire#w2
      I_Contact( "AlarmasDoblePantalla".x40 )
      I_Contact( "AlarmasDoblePantalla".x39 )
      I_Contact( "PanelCompBAJA MTA".MantMC061 )
   END_RUNG wire#w3
   RUNG wire#powerrail
      Contact( "CmpBajaAuto".AutoArrEfMC061 )
      Contact( "CmpBajaAuto".AutoMC061 )
      Contact( "PanelCompBAJA MTA".HabMC061 )
   END_RUNG wire#w2
   RUNG wire#powerrail
      I_Contact( "PanelCompBAJA MTA".InhMC061 )
      I_Contact( "PanelCompBAJA MTA".MantMC061 )
   END_RUNG wire#w4
   // the same network as SCL:
   "MC061 - Compresor de Baja SULLAIR 1"(GMT := "MC061-TO",   // "FB_CTR_MOT"
                           CNF_MAR_D := "MC061-CO" AND NOT "PanelCompBAJA MTA".MantMC061,
                           ORD_MAR_D := (("PanelCompBAJA MTA".MarchaMC061 AND NOT "CmpBajaAuto".AutoMC061) OR ("CmpBajaAuto".AutoArrEfMC061 AND "CmpBajaAuto".AutoMC061 AND "PanelCompBAJA MTA".HabMC061)) AND NOT "AlarmasDoblePantalla".x40 AND NOT "AlarmasDoblePantalla".x39 AND NOT "PanelCompBAJA MTA".MantMC061,
                           MAR_SOLA := "UNO",
                           HAB_ARR_D := NOT "PanelCompBAJA MTA".InhMC061 AND NOT "PanelCompBAJA MTA".MantMC061,
                           INH_MAR_D := "PanelCompBAJA MTA".InhMC061,
                           ACT_MAR_D => "MC061_MARCHA",
                           F_GMT => "DB_ALA_PRE".x39,
                           F_CTC_MAR_D => "DB_ALA_PRE".x40);
END_REGION

REGION Network 18
   RUNG wire#powerrail
      Contact( "MC001" )
      P_Trig( "FlaAuxB1" )
      S_PULSE(T_NO := "ArrMC061", TV := S5T#20S, R :=, BI =>, RET_VAL =>)
      Coil( #TEMP0 )
   END_RUNG
   // the same network as SCL:
   #_w1 := "MC001" AND NOT "FlaAuxB1";   // rising edge
   "FlaAuxB1" := "MC001";
   #_s5time1 := S_PULSE(T_NO := "ArrMC061", S := #_w1, TV := S5T#20S, Q => #_w2);
   #TEMP0 := #_w2;
END_REGION

REGION Network 19: M COMPR BAJA SULLAIR 0-ORDEN PARADA / Parada MC062
   RUNG wire#powerrail
      Contact( "PanelCompBAJA MTA".ParadaPanelMC062 )
      Coil( "Parada-MC062" )
   END_RUNG
   // the same network as SCL:
   "Parada-MC062" := "PanelCompBAJA MTA".ParadaPanelMC062;
END_REGION

REGION Network 20: Motor MC062 - Compresor de Baja SULLAIR 0 / Bloque motor MC062 - Compresor de Baja SULLAIR 0